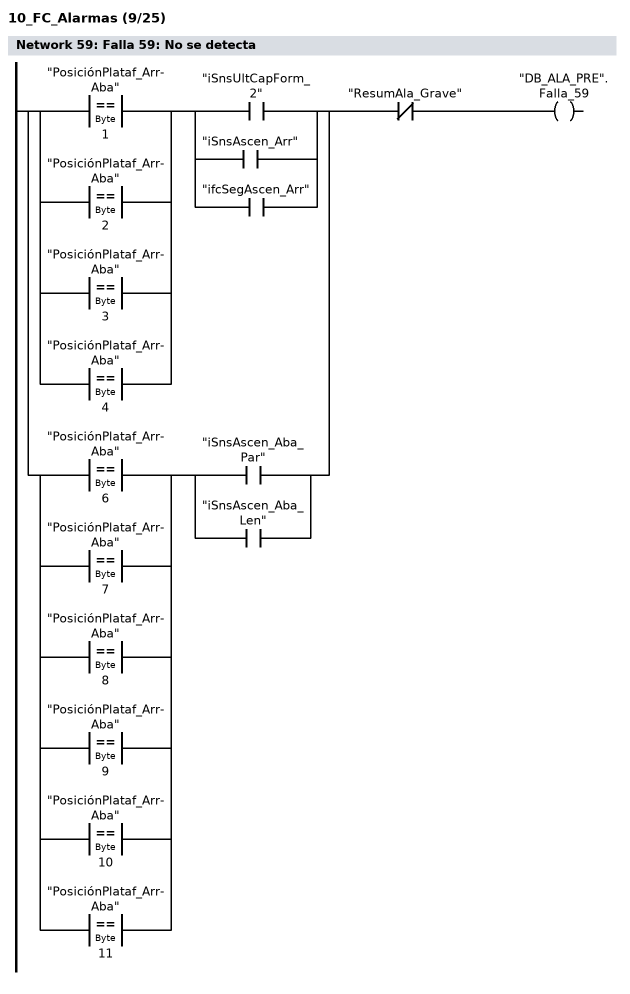
   RUNG wire#powerrail
      { S7_Templates := "SrcType := Byte" } EQ_Contact(in1 := "PosiciónPlataf_Arr-Aba", in2 := 1)
      wire#w1
      Contact( "iSnsUltCapForm_2" )
      wire#w2
      I_Contact( "ResumAla_Grave" )
      Coil( "DB_ALA_PRE".Falla_59 )
   END_RUNG
   RUNG wire#powerrail
      { S7_Templates := "SrcType := Byte" } EQ_Contact(in1 := "PosiciónPlataf_Arr-Aba", in2 := 2)
   END_RUNG wire#w1
   RUNG wire#powerrail
      { S7_Templates := "SrcType := Byte" } EQ_Contact(in1 := "PosiciónPlataf_Arr-Aba", in2 := 3)
   END_RUNG wire#w1
   RUNG wire#powerrail
      { S7_Templates := "SrcType := Byte" } EQ_Contact(in1 := "PosiciónPlataf_Arr-Aba", in2 := 4)
   END_RUNG wire#w1
   RUNG wire#w1
      Contact( "iSnsAscen_Arr" )
   END_RUNG wire#w2
   RUNG wire#w1
      Contact( "ifcSegAscen_Arr" )
   END_RUNG wire#w2
   RUNG wire#powerrail
      { S7_Templates := "SrcType := Byte" } EQ_Contact(in1 := "PosiciónPlataf_Arr-Aba", in2 := 6)
      wire#w3
      Contact( "iSnsAscen_Aba_Par" )
   END_RUNG wire#w2
   RUNG wire#powerrail
      { S7_Templates := "SrcType := Byte" } EQ_Contact(in1 := "PosiciónPlataf_Arr-Aba", in2 := 7)
   END_RUNG wire#w3
   RUNG wire#powerrail
      { S7_Templates := "SrcType := Byte" } EQ_Contact(in1 := "PosiciónPlataf_Arr-Aba", in2 := 8)
   END_RUNG wire#w3
   RUNG wire#powerrail
      { S7_Templates := "SrcType := Byte" } EQ_Contact(in1 := "PosiciónPlataf_Arr-Aba", in2 := 9)
   END_RUNG wire#w3
   RUNG wire#powerrail
      { S7_Templates := "SrcType := Byte" } EQ_Contact(in1 := "PosiciónPlataf_Arr-Aba", in2 := 10)
   END_RUNG wire#w3
   RUNG wire#powerrail
      { S7_Templates := "SrcType := Byte" } EQ_Contact(in1 := "PosiciónPlataf_Arr-Aba", in2 := 11)
   END_RUNG wire#w3
   RUNG wire#w3
      Contact( "iSnsAscen_Aba_Len" )
   END_RUNG wire#w2
   // the same network as SCL:
   "DB_ALA_PRE".Falla_59 := (((("PosiciónPlataf_Arr-Aba" = 1) OR ("PosiciónPlataf_Arr-Aba" = 2) OR ("PosiciónPlataf_Arr-Aba" = 3) OR ("PosiciónPlataf_Arr-Aba" = 4)) AND ("iSnsUltCapForm_2" OR "iSnsAscen_Arr" OR "ifcSegAscen_Arr")) OR ((("PosiciónPlataf_Arr-Aba" = 6) OR ("PosiciónPlataf_Arr-Aba" = 7) OR ("PosiciónPlataf_Arr-Aba" = 8) OR ("PosiciónPlataf_Arr-Aba" = 9) OR ("PosiciónPlataf_Arr-Aba" = 10) OR ("PosiciónPlataf_Arr-Aba" = 11)) AND ("iSnsAscen_Aba_Par" OR "iSnsAscen_Aba_Len"))) AND NOT "ResumAla_Grave";
END_REGION

REGION Network 60: Falla 60: No se detecta
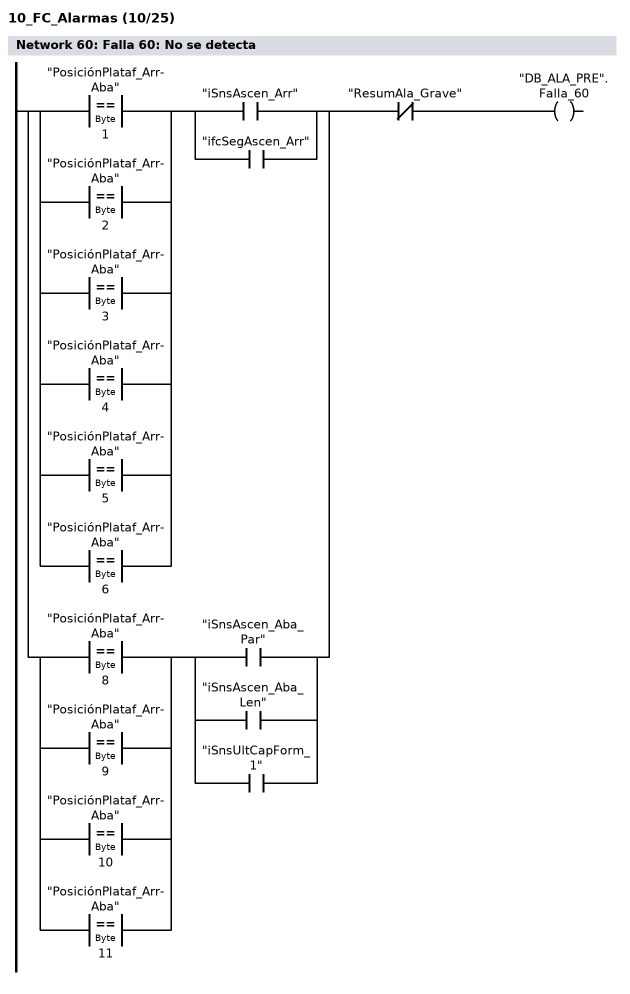
   RUNG wire#powerrail
      { S7_Templates := "SrcType := Byte" } EQ_Contact(in1 := "PosiciónPlataf_Arr-Aba", in2 := 1)
      wire#w1
      Contact( "iSnsAscen_Arr" )
      wire#w2
      I_Contact( "ResumAla_Grave" )
      Coil( "DB_ALA_PRE".Falla_60 )
   END_RUNG
   RUNG wire#powerrail
      { S7_Templates := "SrcType := Byte" } EQ_Contact(in1 := "PosiciónPlataf_Arr-Aba", in2 := 2)
   END_RUNG wire#w1
   RUNG wire#powerrail
      { S7_Templates := "SrcType := Byte" } EQ_Contact(in1 := "PosiciónPlataf_Arr-Aba", in2 := 3)
   END_RUNG wire#w1
   RUNG wire#powerrail
      { S7_Templates := "SrcType := Byte" } EQ_Contact(in1 := "PosiciónPlataf_Arr-Aba", in2 := 4)
   END_RUNG wire#w1
   RUNG wire#powerrail
      { S7_Templates := "SrcType := Byte" } EQ_Contact(in1 := "PosiciónPlataf_Arr-Aba", in2 := 5)
   END_RUNG wire#w1
   RUNG wire#powerrail
      { S7_Templates := "SrcType := Byte" } EQ_Contact(in1 := "PosiciónPlataf_Arr-Aba", in2 := 6)
   END_RUNG wire#w1
   RUNG wire#w1
      Contact( "ifcSegAscen_Arr" )
   END_RUNG wire#w2
   RUNG wire#powerrail
      { S7_Templates := "SrcType := Byte" } EQ_Contact(in1 := "PosiciónPlataf_Arr-Aba", in2 := 8)
      wire#w3
      Contact( "iSnsAscen_Aba_Par" )
   END_RUNG wire#w2
   RUNG wire#powerrail
      { S7_Templates := "SrcType := Byte" } EQ_Contact(in1 := "PosiciónPlataf_Arr-Aba", in2 := 9)
   END_RUNG wire#w3
   RUNG wire#powerrail
      { S7_Templates := "SrcType := Byte" } EQ_Contact(in1 := "PosiciónPlataf_Arr-Aba", in2 := 10)
   END_RUNG wire#w3
   RUNG wire#powerrail
      { S7_Templates := "SrcType := Byte" } EQ_Contact(in1 := "PosiciónPlataf_Arr-Aba", in2 := 11)
   END_RUNG wire#w3
   RUNG wire#w3
      Contact( "iSnsAscen_Aba_Len" )
   END_RUNG wire#w2
   RUNG wire#w3
      Contact( "iSnsUltCapForm_1" )
   END_RUNG wire#w2
   // the same network as SCL:
   "DB_ALA_PRE".Falla_60 := (((("PosiciónPlataf_Arr-Aba" = 1) OR ("PosiciónPlataf_Arr-Aba" = 2) OR ("PosiciónPlataf_Arr-Aba" = 3) OR ("PosiciónPlataf_Arr-Aba" = 4) OR ("PosiciónPlataf_Arr-Aba" = 5) OR ("PosiciónPlataf_Arr-Aba" = 6)) AND ("iSnsAscen_Arr" OR "ifcSegAscen_Arr")) OR ((("PosiciónPlataf_Arr-Aba" = 8) OR ("PosiciónPlataf_Arr-Aba" = 9) OR ("PosiciónPlataf_Arr-Aba" = 10) OR ("PosiciónPlataf_Arr-Aba" = 11)) AND ("iSnsAscen_Aba_Par" OR "iSnsAscen_Aba_Len" OR "iSnsUltCapForm_1"))) AND NOT "ResumAla_Grave";
END_REGION

REGION Network 61: Falla 61: No se detecta Elevador Arriba
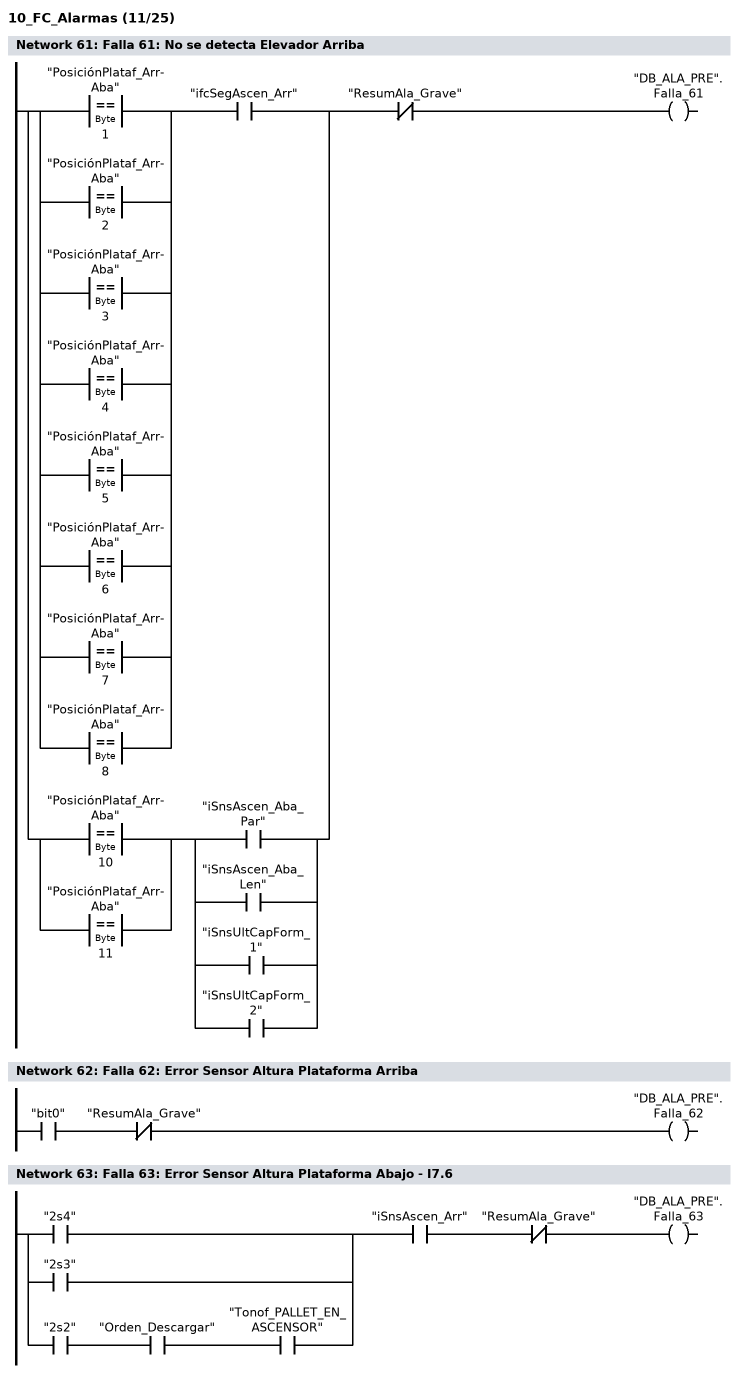
   RUNG wire#powerrail
      { S7_Templates := "SrcType := Byte" } EQ_Contact(in1 := "PosiciónPlataf_Arr-Aba", in2 := 1)
      wire#w1
      Contact( "ifcSegAscen_Arr" )
      wire#w2
      I_Contact( "ResumAla_Grave" )
      Coil( "DB_ALA_PRE".Falla_61 )
   END_RUNG
   RUNG wire#powerrail
      { S7_Templates := "SrcType := Byte" } EQ_Contact(in1 := "PosiciónPlataf_Arr-Aba", in2 := 2)
   END_RUNG wire#w1
   RUNG wire#powerrail
      { S7_Templates := "SrcType := Byte" } EQ_Contact(in1 := "PosiciónPlataf_Arr-Aba", in2 := 3)
   END_RUNG wire#w1
   RUNG wire#powerrail
      { S7_Templates := "SrcType := Byte" } EQ_Contact(in1 := "PosiciónPlataf_Arr-Aba", in2 := 4)
   END_RUNG wire#w1
   RUNG wire#powerrail
      { S7_Templates := "SrcType := Byte" } EQ_Contact(in1 := "PosiciónPlataf_Arr-Aba", in2 := 5)
   END_RUNG wire#w1
   RUNG wire#powerrail
      { S7_Templates := "SrcType := Byte" } EQ_Contact(in1 := "PosiciónPlataf_Arr-Aba", in2 := 6)
   END_RUNG wire#w1
   RUNG wire#powerrail
      { S7_Templates := "SrcType := Byte" } EQ_Contact(in1 := "PosiciónPlataf_Arr-Aba", in2 := 7)
   END_RUNG wire#w1
   RUNG wire#powerrail
      { S7_Templates := "SrcType := Byte" } EQ_Contact(in1 := "PosiciónPlataf_Arr-Aba", in2 := 8)
   END_RUNG wire#w1
   RUNG wire#powerrail
      { S7_Templates := "SrcType := Byte" } EQ_Contact(in1 := "PosiciónPlataf_Arr-Aba", in2 := 10)
      wire#w3
      Contact( "iSnsAscen_Aba_Par" )
   END_RUNG wire#w2
   RUNG wire#powerrail
      { S7_Templates := "SrcType := Byte" } EQ_Contact(in1 := "PosiciónPlataf_Arr-Aba", in2 := 11)
   END_RUNG wire#w3
   RUNG wire#w3
      Contact( "iSnsAscen_Aba_Len" )
   END_RUNG wire#w2
   RUNG wire#w3
      Contact( "iSnsUltCapForm_1" )
   END_RUNG wire#w2
   RUNG wire#w3
      Contact( "iSnsUltCapForm_2" )
   END_RUNG wire#w2
   // the same network as SCL:
   "DB_ALA_PRE".Falla_61 := (((("PosiciónPlataf_Arr-Aba" = 1) OR ("PosiciónPlataf_Arr-Aba" = 2) OR ("PosiciónPlataf_Arr-Aba" = 3) OR ("PosiciónPlataf_Arr-Aba" = 4) OR ("PosiciónPlataf_Arr-Aba" = 5) OR ("PosiciónPlataf_Arr-Aba" = 6) OR ("PosiciónPlataf_Arr-Aba" = 7) OR ("PosiciónPlataf_Arr-Aba" = 8)) AND "ifcSegAscen_Arr") OR ((("PosiciónPlataf_Arr-Aba" = 10) OR ("PosiciónPlataf_Arr-Aba" = 11)) AND ("iSnsAscen_Aba_Par" OR "iSnsAscen_Aba_Len" OR "iSnsUltCapForm_1" OR "iSnsUltCapForm_2"))) AND NOT "ResumAla_Grave";
END_REGION

REGION Network 62: Falla 62: Error Sensor Altura Plataforma Arriba
   RUNG wire#powerrail
      Contact( "bit0" )
      I_Contact( "ResumAla_Grave" )
      Coil( "DB_ALA_PRE".Falla_62 )
   END_RUNG
   // the same network as SCL:
   "DB_ALA_PRE".Falla_62 := "bit0" AND NOT "ResumAla_Grave";
END_REGION

REGION Network 63: Falla 63: Error Sensor Altura Plataforma Abajo - I7.6
   RUNG wire#powerrail
      Contact( "2s4" )
      wire#w1
      Contact( "iSnsAscen_Arr" )
      I_Contact( "ResumAla_Grave" )
      Coil( "DB_ALA_PRE".Falla_63 )
   END_RUNG
   RUNG wire#powerrail
      Contact( "2s3" )
   END_RUNG wire#w1
   RUNG wire#powerrail
      Contact( "2s2" )
      Contact( "Orden_Descargar" )
      Contact( "Tonof_PALLET_EN_ASCENSOR" )
   END_RUNG wire#w1
   // the same network as SCL:
   "DB_ALA_PRE".Falla_63 := ("2s4" OR "2s3" OR ("2s2" AND "Orden_Descargar" AND "Tonof_PALLET_EN_ASCENSOR")) AND "iSnsAscen_Arr" AND NOT "ResumAla_Grave";
END_REGION

REGION Network 64: Falla 64: Error Sensores Altura Plataforma
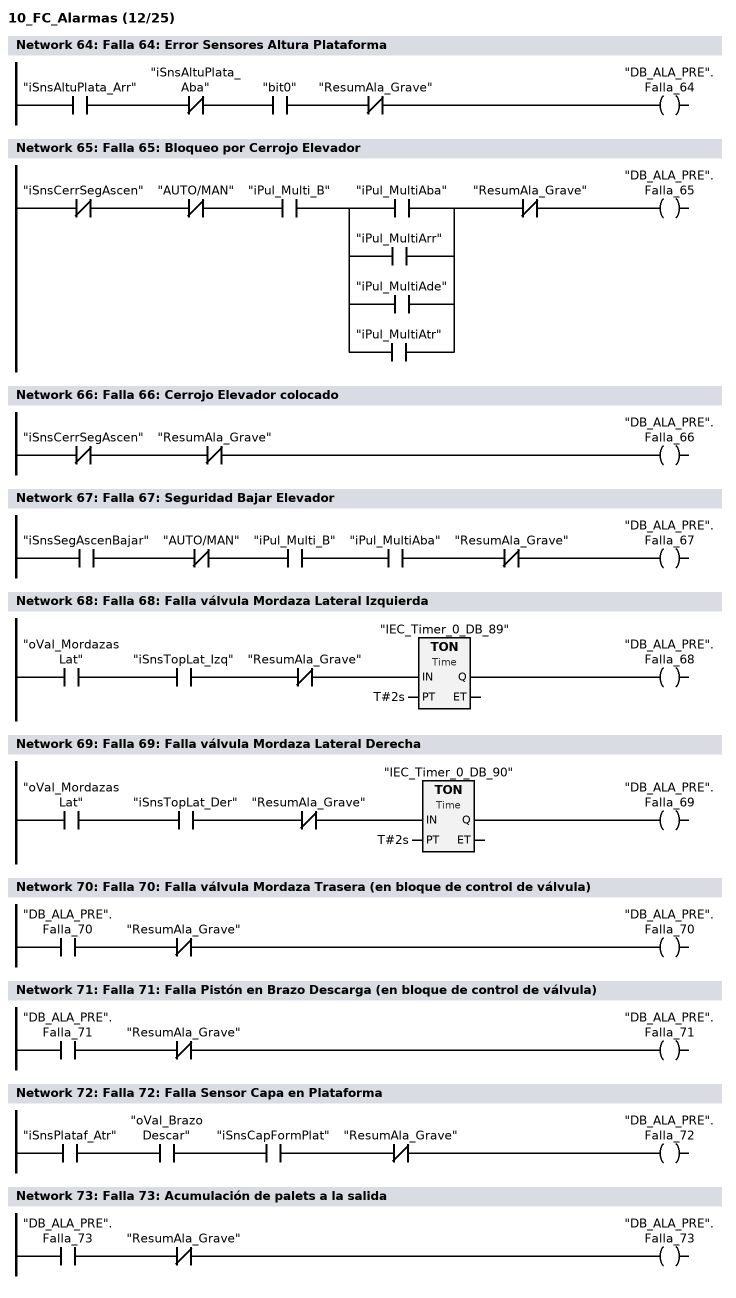
   RUNG wire#powerrail
      Contact( "iSnsAltuPlata_Arr" )
      I_Contact( "iSnsAltuPlata_Aba" )
      Contact( "bit0" )
      I_Contact( "ResumAla_Grave" )
      Coil( "DB_ALA_PRE".Falla_64 )
   END_RUNG
   // the same network as SCL:
   "DB_ALA_PRE".Falla_64 := "iSnsAltuPlata_Arr" AND NOT "iSnsAltuPlata_Aba" AND "bit0" AND NOT "ResumAla_Grave";
END_REGION

REGION Network 65: Falla 65: Bloqueo por Cerrojo Elevador
   RUNG wire#powerrail
      I_Contact( "iSnsCerrSegAscen" )
      I_Contact( "AUTO/MAN" )
      Contact( "iPul_Multi_B" )
      wire#w1
      Contact( "iPul_MultiAba" )
      wire#w2
      I_Contact( "ResumAla_Grave" )
      Coil( "DB_ALA_PRE".Falla_65 )
   END_RUNG
   RUNG wire#w1
      Contact( "iPul_MultiArr" )
   END_RUNG wire#w2
   RUNG wire#w1
      Contact( "iPul_MultiAde" )
   END_RUNG wire#w2
   RUNG wire#w1
      Contact( "iPul_MultiAtr" )
   END_RUNG wire#w2
   // the same network as SCL:
   "DB_ALA_PRE".Falla_65 := NOT "iSnsCerrSegAscen" AND NOT "AUTO/MAN" AND "iPul_Multi_B" AND ("iPul_MultiAba" OR "iPul_MultiArr" OR "iPul_MultiAde" OR "iPul_MultiAtr") AND NOT "ResumAla_Grave";
END_REGION

REGION Network 66: Falla 66: Cerrojo Elevador colocado
   RUNG wire#powerrail
      I_Contact( "iSnsCerrSegAscen" )
      I_Contact( "ResumAla_Grave" )
      Coil( "DB_ALA_PRE".Falla_66 )
   END_RUNG
   // the same network as SCL:
   "DB_ALA_PRE".Falla_66 := NOT "iSnsCerrSegAscen" AND NOT "ResumAla_Grave";
END_REGION

REGION Network 67: Falla 67: Seguridad Bajar Elevador
   RUNG wire#powerrail
      Contact( "iSnsSegAscenBajar" )
      I_Contact( "AUTO/MAN" )
      Contact( "iPul_Multi_B" )
      Contact( "iPul_MultiAba" )
      I_Contact( "ResumAla_Grave" )
      Coil( "DB_ALA_PRE".Falla_67 )
   END_RUNG
   // the same network as SCL:
   "DB_ALA_PRE".Falla_67 := "iSnsSegAscenBajar" AND NOT "AUTO/MAN" AND "iPul_Multi_B" AND "iPul_MultiAba" AND NOT "ResumAla_Grave";
END_REGION

REGION Network 68: Falla 68: Falla válvula Mordaza Lateral Izquierda
   "IEC_Timer_0_DB_89".TON(IN := "oVal_MordazasLat" AND "iSnsTopLat_Izq" AND NOT "ResumAla_Grave", PT := T#2s);
   "DB_ALA_PRE".Falla_68 := "IEC_Timer_0_DB_89".Q;
END_REGION

REGION Network 69: Falla 69: Falla válvula Mordaza Lateral Derecha
   "IEC_Timer_0_DB_90".TON(IN := "oVal_MordazasLat" AND "iSnsTopLat_Der" AND NOT "ResumAla_Grave", PT := T#2s);
   "DB_ALA_PRE".Falla_69 := "IEC_Timer_0_DB_90".Q;
END_REGION

REGION Network 70: Falla 70: Falla válvula Mordaza Trasera (en bloque de control de válvula)
   RUNG wire#powerrail
      Contact( "DB_ALA_PRE".Falla_70 )
      I_Contact( "ResumAla_Grave" )
      Coil( "DB_ALA_PRE".Falla_70 )
   END_RUNG
   // the same network as SCL:
   "DB_ALA_PRE".Falla_70 := "DB_ALA_PRE".Falla_70 AND NOT "ResumAla_Grave";
END_REGION

REGION Network 71: Falla 71: Falla Pistón en Brazo Descarga (en bloque de control de válvula)
   RUNG wire#powerrail
      Contact( "DB_ALA_PRE".Falla_71 )
      I_Contact( "ResumAla_Grave" )
      Coil( "DB_ALA_PRE".Falla_71 )
   END_RUNG
   // the same network as SCL:
   "DB_ALA_PRE".Falla_71 := "DB_ALA_PRE".Falla_71 AND NOT "ResumAla_Grave";
END_REGION

REGION Network 72: Falla 72: Falla Sensor Capa en Plataforma
   RUNG wire#powerrail
      Contact( "iSnsPlataf_Atr" )
      Contact( "oVal_BrazoDescar" )
      Contact( "iSnsCapFormPlat" )
      I_Contact( "ResumAla_Grave" )
      Coil( "DB_ALA_PRE".Falla_72 )
   END_RUNG
   // the same network as SCL:
   "DB_ALA_PRE".Falla_72 := "iSnsPlataf_Atr" AND "oVal_BrazoDescar" AND "iSnsCapFormPlat" AND NOT "ResumAla_Grave";
END_REGION

REGION Network 73: Falla 73: Acumulación de palets a la salida
   RUNG wire#powerrail
      Contact( "DB_ALA_PRE".Falla_73 )
      I_Contact( "ResumAla_Grave" )
      Coil( "DB_ALA_PRE".Falla_73 )
   END_RUNG
   // the same network as SCL:
   "DB_ALA_PRE".Falla_73 := "DB_ALA_PRE".Falla_73 AND NOT "ResumAla_Grave";
END_REGION

REGION Network 74: Falla 74:
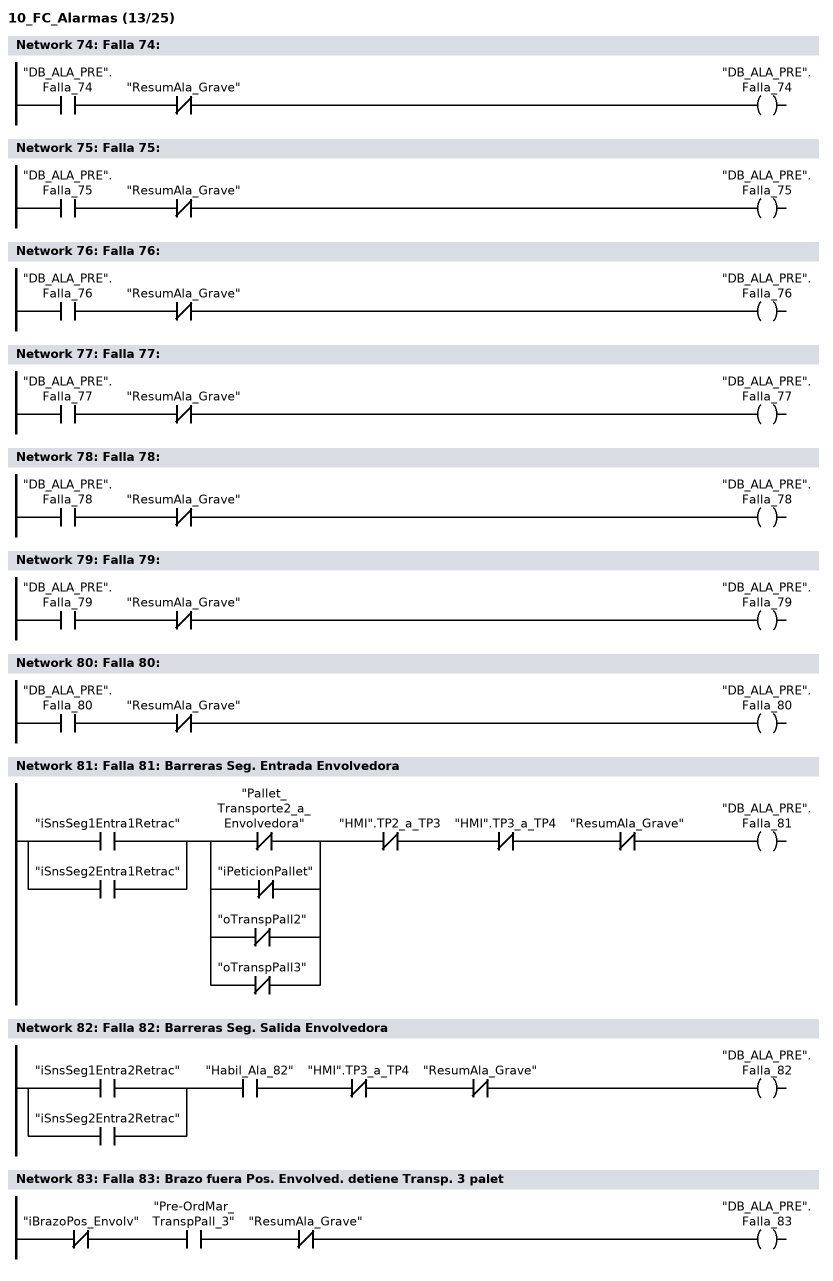
   RUNG wire#powerrail
      Contact( "DB_ALA_PRE".Falla_74 )
      I_Contact( "ResumAla_Grave" )
      Coil( "DB_ALA_PRE".Falla_74 )
   END_RUNG
   // the same network as SCL:
   "DB_ALA_PRE".Falla_74 := "DB_ALA_PRE".Falla_74 AND NOT "ResumAla_Grave";
END_REGION

REGION Network 75: Falla 75:
   RUNG wire#powerrail
      Contact( "DB_ALA_PRE".Falla_75 )
      I_Contact( "ResumAla_Grave" )
      Coil( "DB_ALA_PRE".Falla_75 )
   END_RUNG
   // the same network as SCL:
   "DB_ALA_PRE".Falla_75 := "DB_ALA_PRE".Falla_75 AND NOT "ResumAla_Grave";
END_REGION

REGION Network 76: Falla 76:
   RUNG wire#powerrail
      Contact( "DB_ALA_PRE".Falla_76 )
      I_Contact( "ResumAla_Grave" )
      Coil( "DB_ALA_PRE".Falla_76 )
   END_RUNG
   // the same network as SCL:
   "DB_ALA_PRE".Falla_76 := "DB_ALA_PRE".Falla_76 AND NOT "ResumAla_Grave";
END_REGION

REGION Network 77: Falla 77:
   RUNG wire#powerrail
      Contact( "DB_ALA_PRE".Falla_77 )
      I_Contact( "ResumAla_Grave" )
      Coil( "DB_ALA_PRE".Falla_77 )
   END_RUNG
   // the same network as SCL:
   "DB_ALA_PRE".Falla_77 := "DB_ALA_PRE".Falla_77 AND NOT "ResumAla_Grave";
END_REGION

REGION Network 78: Falla 78:
   RUNG wire#powerrail
      Contact( "DB_ALA_PRE".Falla_78 )
      I_Contact( "ResumAla_Grave" )
      Coil( "DB_ALA_PRE".Falla_78 )
   END_RUNG
   // the same network as SCL:
   "DB_ALA_PRE".Falla_78 := "DB_ALA_PRE".Falla_78 AND NOT "ResumAla_Grave";
END_REGION

REGION Network 79: Falla 79:
   RUNG wire#powerrail
      Contact( "DB_ALA_PRE".Falla_79 )
      I_Contact( "ResumAla_Grave" )
      Coil( "DB_ALA_PRE".Falla_79 )
   END_RUNG
   // the same network as SCL:
   "DB_ALA_PRE".Falla_79 := "DB_ALA_PRE".Falla_79 AND NOT "ResumAla_Grave";
END_REGION

REGION Network 80: Falla 80:
   RUNG wire#powerrail
      Contact( "DB_ALA_PRE".Falla_80 )
      I_Contact( "ResumAla_Grave" )
      Coil( "DB_ALA_PRE".Falla_80 )
   END_RUNG
   // the same network as SCL:
   "DB_ALA_PRE".Falla_80 := "DB_ALA_PRE".Falla_80 AND NOT "ResumAla_Grave";
END_REGION

REGION Network 81: Falla 81: Barreras Seg. Entrada Envolvedora
   RUNG wire#powerrail
      Contact( "iSnsSeg1Entra1Retrac" )
      wire#w1
      I_Contact( "Pallet_Transporte2_a_Envolvedora" )
      wire#w2
      I_Contact( "HMI".TP2_a_TP3 )
      I_Contact( "HMI".TP3_a_TP4 )
      I_Contact( "ResumAla_Grave" )
      Coil( "DB_ALA_PRE".Falla_81 )
   END_RUNG
   RUNG wire#powerrail
      Contact( "iSnsSeg2Entra1Retrac" )
   END_RUNG wire#w1
   RUNG wire#w1
      I_Contact( "iPeticionPallet" )
   END_RUNG wire#w2
   RUNG wire#w1
      I_Contact( "oTranspPall2" )
   END_RUNG wire#w2
   RUNG wire#w1
      I_Contact( "oTranspPall3" )
   END_RUNG wire#w2
   // the same network as SCL:
   "DB_ALA_PRE".Falla_81 := ("iSnsSeg1Entra1Retrac" OR "iSnsSeg2Entra1Retrac") AND (NOT "Pallet_Transporte2_a_Envolvedora" OR NOT "iPeticionPallet" OR NOT "oTranspPall2" OR NOT "oTranspPall3") AND NOT "HMI".TP2_a_TP3 AND NOT "HMI".TP3_a_TP4 AND NOT "ResumAla_Grave";
END_REGION

REGION Network 82: Falla 82: Barreras Seg. Salida Envolvedora
   RUNG wire#powerrail
      Contact( "iSnsSeg1Entra2Retrac" )
      wire#w1
      Contact( "Habil_Ala_82" )
      I_Contact( "HMI".TP3_a_TP4 )
      I_Contact( "ResumAla_Grave" )
      Coil( "DB_ALA_PRE".Falla_82 )
   END_RUNG
   RUNG wire#powerrail
      Contact( "iSnsSeg2Entra2Retrac" )
   END_RUNG wire#w1
   // the same network as SCL:
   "DB_ALA_PRE".Falla_82 := ("iSnsSeg1Entra2Retrac" OR "iSnsSeg2Entra2Retrac") AND "Habil_Ala_82" AND NOT "HMI".TP3_a_TP4 AND NOT "ResumAla_Grave";
END_REGION

REGION Network 83: Falla 83: Brazo fuera Pos. Envolved. detiene Transp. 3 palet
   RUNG wire#powerrail
      I_Contact( "iBrazoPos_Envolv" )
      Contact( "Pre-OrdMar_TranspPall_3" )
      I_Contact( "ResumAla_Grave" )
      Coil( "DB_ALA_PRE".Falla_83 )
   END_RUNG
   // the same network as SCL:
   "DB_ALA_PRE".Falla_83 := NOT "iBrazoPos_Envolv" AND "Pre-OrdMar_TranspPall_3" AND NOT "ResumAla_Grave";
END_REGION

REGION Network 84: Falla 84:
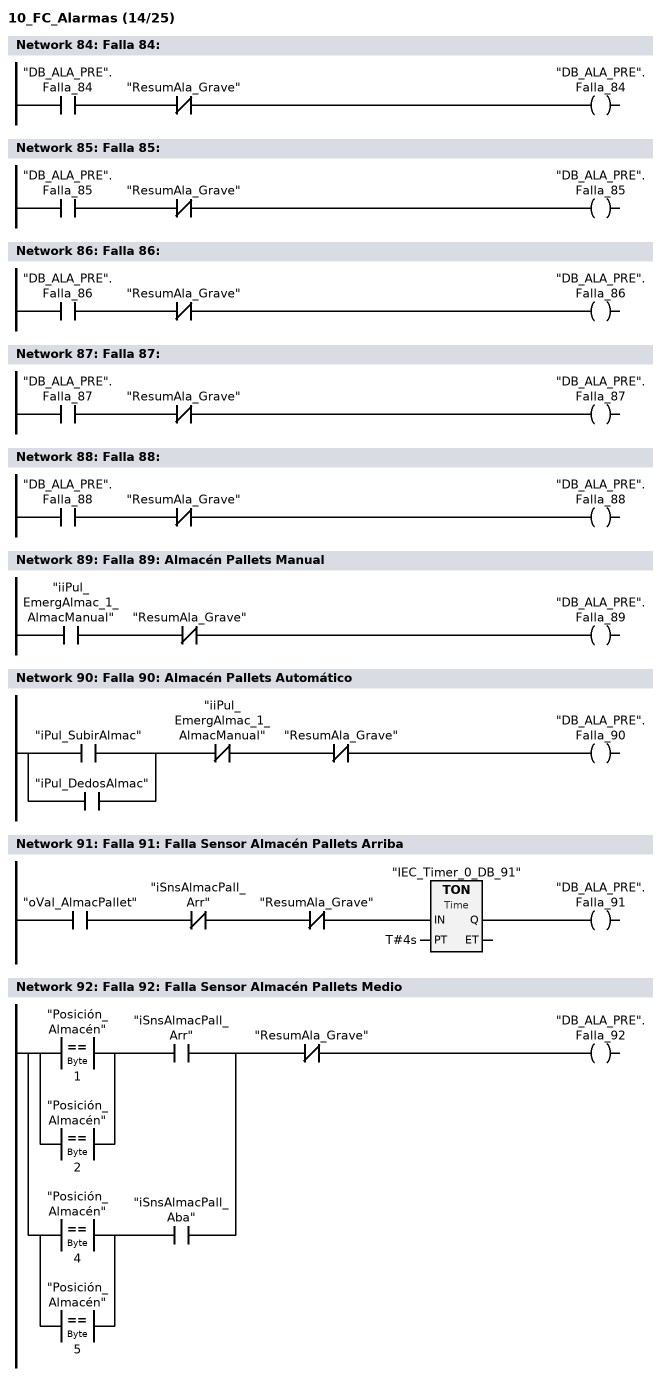
   RUNG wire#powerrail
      Contact( "DB_ALA_PRE".Falla_84 )
      I_Contact( "ResumAla_Grave" )
      Coil( "DB_ALA_PRE".Falla_84 )
   END_RUNG
   // the same network as SCL:
   "DB_ALA_PRE".Falla_84 := "DB_ALA_PRE".Falla_84 AND NOT "ResumAla_Grave";
END_REGION

REGION Network 85: Falla 85:
   RUNG wire#powerrail
      Contact( "DB_ALA_PRE".Falla_85 )
      I_Contact( "ResumAla_Grave" )
      Coil( "DB_ALA_PRE".Falla_85 )
   END_RUNG
   // the same network as SCL:
   "DB_ALA_PRE".Falla_85 := "DB_ALA_PRE".Falla_85 AND NOT "ResumAla_Grave";
END_REGION

REGION Network 86: Falla 86:
   RUNG wire#powerrail
      Contact( "DB_ALA_PRE".Falla_86 )
      I_Contact( "ResumAla_Grave" )
      Coil( "DB_ALA_PRE".Falla_86 )
   END_RUNG
   // the same network as SCL:
   "DB_ALA_PRE".Falla_86 := "DB_ALA_PRE".Falla_86 AND NOT "ResumAla_Grave";
END_REGION

REGION Network 87: Falla 87:
   RUNG wire#powerrail
      Contact( "DB_ALA_PRE".Falla_87 )
      I_Contact( "ResumAla_Grave" )
      Coil( "DB_ALA_PRE".Falla_87 )
   END_RUNG
   // the same network as SCL:
   "DB_ALA_PRE".Falla_87 := "DB_ALA_PRE".Falla_87 AND NOT "ResumAla_Grave";
END_REGION

REGION Network 88: Falla 88:
   RUNG wire#powerrail
      Contact( "DB_ALA_PRE".Falla_88 )
      I_Contact( "ResumAla_Grave" )
      Coil( "DB_ALA_PRE".Falla_88 )
   END_RUNG
   // the same network as SCL:
   "DB_ALA_PRE".Falla_88 := "DB_ALA_PRE".Falla_88 AND NOT "ResumAla_Grave";
END_REGION

REGION Network 89: Falla 89: Almacén Pallets Manual
   RUNG wire#powerrail
      Contact( "iiPul_EmergAlmac_1_AlmacManual" )
      I_Contact( "ResumAla_Grave" )
      Coil( "DB_ALA_PRE".Falla_89 )
   END_RUNG
   // the same network as SCL:
   "DB_ALA_PRE".Falla_89 := "iiPul_EmergAlmac_1_AlmacManual" AND NOT "ResumAla_Grave";
END_REGION

REGION Network 90: Falla 90: Almacén Pallets Automático
   RUNG wire#powerrail
      Contact( "iPul_SubirAlmac" )
      wire#w1
      I_Contact( "iiPul_EmergAlmac_1_AlmacManual" )
      I_Contact( "ResumAla_Grave" )
      Coil( "DB_ALA_PRE".Falla_90 )
   END_RUNG
   RUNG wire#powerrail
      Contact( "iPul_DedosAlmac" )
   END_RUNG wire#w1
   // the same network as SCL:
   "DB_ALA_PRE".Falla_90 := ("iPul_SubirAlmac" OR "iPul_DedosAlmac") AND NOT "iiPul_EmergAlmac_1_AlmacManual" AND NOT "ResumAla_Grave";
END_REGION

REGION Network 91: Falla 91: Falla Sensor Almacén Pallets Arriba
   "IEC_Timer_0_DB_91".TON(IN := "oVal_AlmacPallet" AND NOT "iSnsAlmacPall_Arr" AND NOT "ResumAla_Grave",
                           PT := T#4s);
   "DB_ALA_PRE".Falla_91 := "IEC_Timer_0_DB_91".Q;
END_REGION

REGION Network 92: Falla 92: Falla Sensor Almacén Pallets Medio
   RUNG wire#powerrail
      { S7_Templates := "SrcType := Byte" } EQ_Contact(in1 := "Posición_Almacén", in2 := 1)
      wire#w1
      Contact( "iSnsAlmacPall_Arr" )
      wire#w2
      I_Contact( "ResumAla_Grave" )
      Coil( "DB_ALA_PRE".Falla_92 )
   END_RUNG
   RUNG wire#powerrail
      { S7_Templates := "SrcType := Byte" } EQ_Contact(in1 := "Posición_Almacén", in2 := 2)
   END_RUNG wire#w1
   RUNG wire#powerrail
      { S7_Templates := "SrcType := Byte" } EQ_Contact(in1 := "Posición_Almacén", in2 := 4)
      wire#w3
      Contact( "iSnsAlmacPall_Aba" )
   END_RUNG wire#w2
   RUNG wire#powerrail
      { S7_Templates := "SrcType := Byte" } EQ_Contact(in1 := "Posición_Almacén", in2 := 5)
   END_RUNG wire#w3
   // the same network as SCL:
   "DB_ALA_PRE".Falla_92 := (((("Posición_Almacén" = 1) OR ("Posición_Almacén" = 2)) AND "iSnsAlmacPall_Arr") OR ((("Posición_Almacén" = 4) OR ("Posición_Almacén" = 5)) AND "iSnsAlmacPall_Aba")) AND NOT "ResumAla_Grave";
END_REGION

REGION Network 93: Falla 93: Falla Sensor Almacén Pallets Abajo
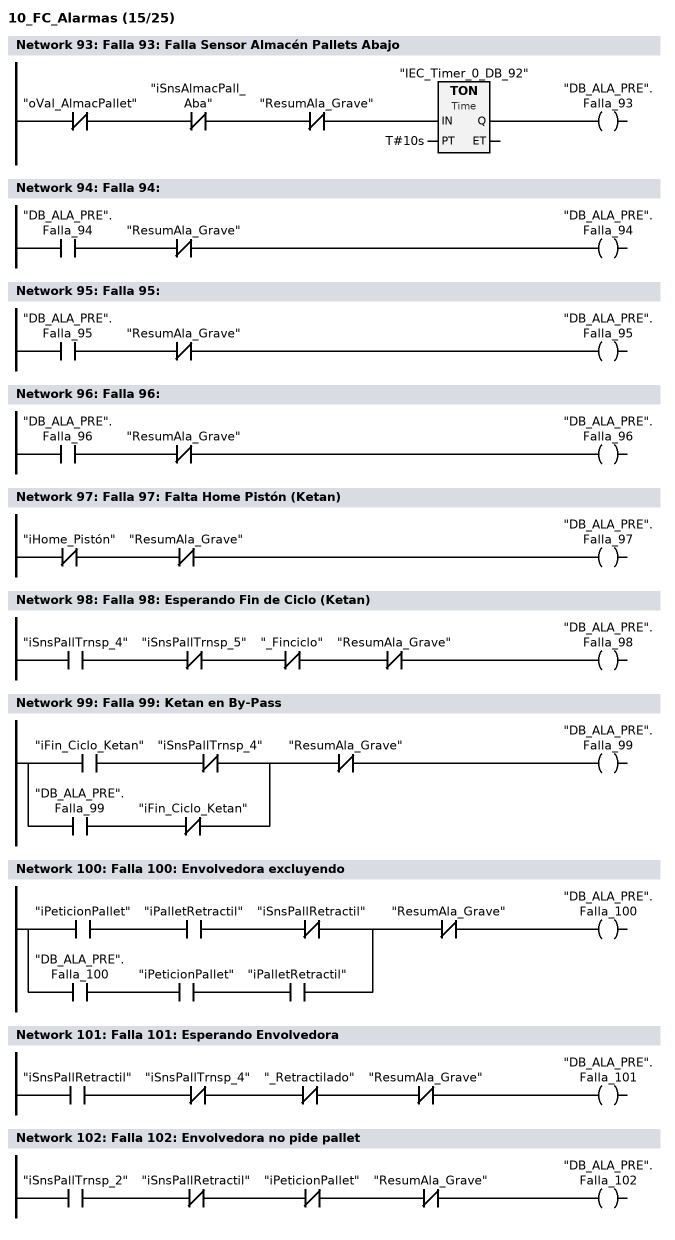
   "IEC_Timer_0_DB_92".TON(IN := NOT "oVal_AlmacPallet" AND NOT "iSnsAlmacPall_Aba" AND NOT "ResumAla_Grave",
                           PT := T#10s);
   "DB_ALA_PRE".Falla_93 := "IEC_Timer_0_DB_92".Q;
END_REGION

REGION Network 94: Falla 94:
   RUNG wire#powerrail
      Contact( "DB_ALA_PRE".Falla_94 )
      I_Contact( "ResumAla_Grave" )
      Coil( "DB_ALA_PRE".Falla_94 )
   END_RUNG
   // the same network as SCL:
   "DB_ALA_PRE".Falla_94 := "DB_ALA_PRE".Falla_94 AND NOT "ResumAla_Grave";
END_REGION

REGION Network 95: Falla 95:
   RUNG wire#powerrail
      Contact( "DB_ALA_PRE".Falla_95 )
      I_Contact( "ResumAla_Grave" )
      Coil( "DB_ALA_PRE".Falla_95 )
   END_RUNG
   // the same network as SCL:
   "DB_ALA_PRE".Falla_95 := "DB_ALA_PRE".Falla_95 AND NOT "ResumAla_Grave";
END_REGION

REGION Network 96: Falla 96:
   RUNG wire#powerrail
      Contact( "DB_ALA_PRE".Falla_96 )
      I_Contact( "ResumAla_Grave" )
      Coil( "DB_ALA_PRE".Falla_96 )
   END_RUNG
   // the same network as SCL:
   "DB_ALA_PRE".Falla_96 := "DB_ALA_PRE".Falla_96 AND NOT "ResumAla_Grave";
END_REGION

REGION Network 97: Falla 97: Falta Home Pistón (Ketan)
   RUNG wire#powerrail
      I_Contact( "iHome_Pistón" )
      I_Contact( "ResumAla_Grave" )
      Coil( "DB_ALA_PRE".Falla_97 )
   END_RUNG
   // the same network as SCL:
   "DB_ALA_PRE".Falla_97 := NOT "iHome_Pistón" AND NOT "ResumAla_Grave";
END_REGION

REGION Network 98: Falla 98: Esperando Fin de Ciclo (Ketan)
   RUNG wire#powerrail
      Contact( "iSnsPallTrnsp_4" )
      I_Contact( "iSnsPallTrnsp_5" )
      I_Contact( "_Finciclo" )
      I_Contact( "ResumAla_Grave" )
      Coil( "DB_ALA_PRE".Falla_98 )
   END_RUNG
   // the same network as SCL:
   "DB_ALA_PRE".Falla_98 := "iSnsPallTrnsp_4" AND NOT "iSnsPallTrnsp_5" AND NOT "_Finciclo" AND NOT "ResumAla_Grave";
END_REGION

REGION Network 99: Falla 99: Ketan en By-Pass
   RUNG wire#powerrail
      Contact( "iFin_Ciclo_Ketan" )
      I_Contact( "iSnsPallTrnsp_4" )
      wire#w1
      I_Contact( "ResumAla_Grave" )
      Coil( "DB_ALA_PRE".Falla_99 )
   END_RUNG
   RUNG wire#powerrail
      Contact( "DB_ALA_PRE".Falla_99 )
      I_Contact( "iFin_Ciclo_Ketan" )
   END_RUNG wire#w1
   // the same network as SCL:
   "DB_ALA_PRE".Falla_99 := (("iFin_Ciclo_Ketan" AND NOT "iSnsPallTrnsp_4") OR ("DB_ALA_PRE".Falla_99 AND NOT "iFin_Ciclo_Ketan")) AND NOT "ResumAla_Grave";
END_REGION

REGION Network 100: Falla 100: Envolvedora excluyendo
   RUNG wire#powerrail
      Contact( "iPeticionPallet" )
      Contact( "iPalletRetractil" )
      I_Contact( "iSnsPallRetractil" )
      wire#w1
      I_Contact( "ResumAla_Grave" )
      Coil( "DB_ALA_PRE".Falla_100 )
   END_RUNG
   RUNG wire#powerrail
      Contact( "DB_ALA_PRE".Falla_100 )
      Contact( "iPeticionPallet" )
      Contact( "iPalletRetractil" )
   END_RUNG wire#w1
   // the same network as SCL:
   "DB_ALA_PRE".Falla_100 := (("iPeticionPallet" AND "iPalletRetractil" AND NOT "iSnsPallRetractil") OR ("DB_ALA_PRE".Falla_100 AND "iPeticionPallet" AND "iPalletRetractil")) AND NOT "ResumAla_Grave";
END_REGION

REGION Network 101: Falla 101: Esperando Envolvedora
   RUNG wire#powerrail
      Contact( "iSnsPallRetractil" )
      I_Contact( "iSnsPallTrnsp_4" )
      I_Contact( "_Retractilado" )
      I_Contact( "ResumAla_Grave" )
      Coil( "DB_ALA_PRE".Falla_101 )
   END_RUNG
   // the same network as SCL:
   "DB_ALA_PRE".Falla_101 := "iSnsPallRetractil" AND NOT "iSnsPallTrnsp_4" AND NOT "_Retractilado" AND NOT "ResumAla_Grave";
END_REGION

REGION Network 102: Falla 102: Envolvedora no pide pallet
   RUNG wire#powerrail
      Contact( "iSnsPallTrnsp_2" )
      I_Contact( "iSnsPallRetractil" )
      I_Contact( "iPeticionPallet" )
      I_Contact( "ResumAla_Grave" )
      Coil( "DB_ALA_PRE".Falla_102 )
   END_RUNG
   // the same network as SCL:
   "DB_ALA_PRE".Falla_102 := "iSnsPallTrnsp_2" AND NOT "iSnsPallRetractil" AND NOT "iPeticionPallet" AND NOT "ResumAla_Grave";
END_REGION

REGION Network 103: Falla 103: No se detecta pallet en Elevador